                 // Copy actual to old
                 #statActualCommandOld := #statActualCommand;
                 #statModalCommandOld := #statModalCommand;

                 // Reset path data element and modal path data element
                 #statActualCommand := #statPathDataElementEmpty;
                 #statModalCommand := #statPathDataElementEmpty;

                 // Reset parameter counter for command
                 #statElementCounter := #statElementCounterEmpty;

                 // Initialize statCompletedPathDataCommand
                 #statActualCommand.pathDataElement := #statPathDataElementEmpty.pathDataElement;

                 FOR #tempCounter := 1 TO "LKINLANG_NUMBER_OF_CONDITIONS" DO
                   #statConditionsToCheck[#tempCounter] := #statConditionEmpty;
                   #statSetParametersInCmd[#tempCounter] := #statConditionEmpty;
                 END_FOR;

                 FOR #tempCounter := 1 TO "LKINLANG_MAX_NUMBER_OF_PARAMETERS_PER_LINE" DO
                   #tempParameterCounter[#tempCounter].parameterNumber := 0;
                   #tempParameterCounter[#tempCounter].counterValue := 0;
                 END_FOR;

                 // Save last positiong state (rel / abs)
                 #statPositioningModeOld := #statPositioningMode;

                 IF #statSearchedLine <= 0 THEN
                   // Next state --> Tokenize new line
                   #statStateIntern := #STATE_TOKENIZING;
                 ELSE
                   // Next state --> Search line
                   #statStateIntern := #STATE_SEARCH_LINE;
                 END_IF;

               END_IF;
             END_REGION RESET_AFTER_WRITE

             // ------------------------------------------------------------------------------------------
             // PreprocessingStop state for internal case
             // Switch to in case of preprocessingStop and do not execute other states
             // Wait until MovePath signalizes done
             // If done then go to STATE_TOKENIZING (continue with next line)
             // ------------------------------------------------------------------------------------------ 
             REGION PREPROCESSING_STOP
               // preprocessingStop State 
               IF #statStateIntern = #STATE_PREPROCESSING_STOP THEN
                 // preprocessingStop bit is set by parser and reset by MovePath 
                 // MovePath resets preprocessingStop if all commands are done
                 // Check if all commands are executed
                 IF #pathData.pointers.preprocessingStop = FALSE THEN
                   // Continue parsing
                   #statStateIntern := #STATE_TOKENIZING;
                 ELSE
                   ; // Stay here and wait
                 END_IF;
               END_IF;
             END_REGION PREPROCESSING_STOP

           END_FOR; // End of for loop 
         END_REGION FB_STATE_PARSING

         // ------------------------------------------------------------------------------------------
         // Error state for internal case
         // Switch to in case of error and do not execute other states
         // ------------------------------------------------------------------------------------------ 
         REGION ERROR_STATE
           // Error State 
           IF #statStateIntern = #STATE_ERROR THEN
             // Reset lineBuffer pointer
             #lineBuffer.pointers.retrievePointer := 0;
             #lineBuffer.pointers.addPointerRestarted := FALSE;
             IF #lineBuffer.pointers.endOfFile = FALSE THEN
               #lineBuffer.pointers.endOfFile := TRUE; // Signalize end to filehandler
             END_IF;
             // Reset file state
             IF #lineBuffer.info.fileState = "LKINLANG_FILE_STATE_RUNNING" THEN
               #lineBuffer.info.fileState := "LKINLANG_FILE_STATE_IDLE";
             END_IF;
           END_IF;
         END_REGION ERROR_STATE


         // ------------------------------------------------------------------------------------------
         // Stopping state in case stop input is triggered
         // Reset pointers where needed
         // ------------------------------------------------------------------------------------------ 
       #FB_STATE_STOPPING: // Stopping the parser
         REGION FB_STATE_STOPPING
           // Reset lineBuffer pointer
           #lineBuffer.pointers.retrievePointer := 0;

           // Reset pathData pointer 
           #pathData.pointers.addPointer := 0;
           #pathData.pointers.ignoreAddPointer := TRUE;
           #pathData.pointers.addPointerRestarted := FALSE;
           #pathData.pointers.bufferLocked := FALSE;
           #pathData.pointers.preprocessingStop := FALSE;

           // Set status
           #statStatus := #STATUS_COMMAND_ABORTED;
         END_REGION FB_STATE_STOPPING

       ELSE // Undefined state in state machine reached
         #statStatus := #ERR_UNDEFINED_STATE;
     END_CASE;

   END_REGION STATE_MACHINE


   REGION OUTPUTS
     // Write outputs
     IF (#statStatus = #STATUS_EXECUTION_FINISHED) AND (#statDone = FALSE) THEN // Execution finished without errors
       #statDone := TRUE;
       #statBusy := FALSE;
       #statCommandAborted := FALSE;
       #statError := FALSE;
       #statFBState := #FB_STATE_NO_PROCESSING; // Switch state machine to "no processing"

     ELSIF (#statStatus.%X15 = TRUE) AND (#statError = FALSE) THEN // Error occurred (#statStatus is 16#8000 to 16#FFFF)
       #statDone := FALSE;
       #statBusy := FALSE;
       #statCommandAborted := FALSE;
       #statError := TRUE;
       #statFBState := #FB_STATE_NO_PROCESSING; // Switch state machine to "no processing"

     ELSIF (#statStatus = #STATUS_COMMAND_ABORTED) AND (#statCommandAborted = FALSE) THEN // Commanded functionality has been aborted by another command
       #statDone := FALSE;
       #statBusy := FALSE;
       #statCommandAborted := TRUE;
       #statError := FALSE;
       #statFBState := #FB_STATE_NO_PROCESSING; // Switch state machine to "no processing"

     ELSIF (#tempExecute = FALSE) AND ((#statDone = TRUE) OR (#statError = TRUE) OR (#statCommandAborted = TRUE)) THEN // Reset outputs
       #statDone := FALSE;
       #statBusy := FALSE;
       #statCommandAborted := FALSE;
       #statError := FALSE;
       #statStatus := #STATUS_NO_CALL;
       // Reset application specific outputs
       #statErrorString := '';
       IF #lineBuffer.info.fileState = "LKINLANG_FILE_STATE_RUNNING" THEN
         #lineBuffer.info.fileState := "LKINLANG_FILE_STATE_IDLE";
       END_IF;
     END_IF;

     // Write static values to outputs
     #done := #statDone;
     #busy := #statBusy;
     #commandAborted := #statCommandAborted;
     #error := #statError;
     #status := #statStatus;
     #errorString := #statErrorString;
   END_REGION OUTPUTS


   //--------------------------------------------------------------------
   // End of Block LKinLang_Parser
   //--------------------------------------------------------------------
END_FUNCTION_BLOCK

FUNCTION_BLOCK "LKinLang_Filehandler"   // FB35451, SCL
TITLE = LKinLang_FileHandler
{ S7_Optimized_Access := 'TRUE' }
AUTHOR : tech.team.motioncontrol@siemens.com
FAMILY : LKinLang
VERSION : 1.1
// Transfer of data between memory card text file and PLC DB (buffer)
   VAR_INPUT
      executePlcToCard : Bool;   // Write data from buffer to card file
      executeCardToPlc : Bool;   // Write data from card file to buffer
      stop : Bool;   // stop the data transfer, abort the current command
      fileName : String;   // name of the card file (e.g. 'ProgramSlot.txt')
   END_VAR
   VAR_OUTPUT
      busy : Bool;   // TRUE: FB is not finished and new output values can be expected
      done : Bool;   // TRUE: Commanded action has been completed successfully
      dataTransferStopped : Bool;   // TRUE: The data transfer has been stopped
      error : Bool;   // Rising edge informs that an error occurred during the execution of
      status : Word := 16#7000;   // Current status of FB
      diagnostics : "LKinLang_typeFileHandlerDiagnostics";   // Diagnostics structure of FB
   END_VAR
   VAR_IN_OUT
      lineBuffer : "LKinLang_typeLineBuffer";   // String buffer connection
   END_VAR
   VAR
      statBusy : Bool;   // Static value for output busy
      statDone : Bool;   // Static value for output done
      statError : Bool;   // Static value for output error
      statCommandAborted : Bool;   // Static value for output commandAborted
      statPlcToCardOld : Bool;   // Old value of execute for edge detection
      statCardToPlcOld : Bool;   // Old value of execute for edge detection
      statStopOld : Bool;   // Old value of stop for edge detection
      statFBState : UInt;   // Static value for FB state
      statByteLine : Array[0..#NUMBER_OF_BYTES_PER_REQUEST] of Byte;   // Data storage for file read/write
      statByteLineCounter : UDInt;   // Counter/Index for the current byte line, which will be written with FileWriteC / Counter in the data storage
      statByteOffsetFile : UDInt;   // Offset for file read/write in the actual file on memory card / Offset for file read/write
      instFileWriteC : FileWriteC;
      instFileReadC : FileReadC;
      statLineCount : UDInt := 0;   // Actual line to write into the DB or into the file on the memory card / Number of lines from the current read file request
      statCurrentByteLine : Array[0..#NUMBER_OF_BYTES_PER_REQUEST] of Byte;   // Read bytes from actual read request
      statCharPosition : DInt;   // Conversion index CHAR-->STRING
      statBufferedLines : Array[0..#MAX_NUMBER_OF_LINES_PER_READ_REQUEST] of "LKinLang_typeLineContent";   // Buffer for single lines of file as string
      statLineIndex : DInt;   // Static store for last written line to continue FOR loop in case of exit
      statLineCountTotal : UDInt;   // Number of lines read in total
      statLastWrittenLine : UDInt;   // Static storing of the last written index
      statReadLineOld : UDInt;   // Static storing of the last read index
      statNumberOfRestBytes : UDInt;   // Number of bytes to be written on to the card
      statFileName : String;   // Static storing for the fileName input
      statFolderName : String := 'UserFiles';   // Static storing for the folderName
      statStatus : Word := 16#7000;   // Static value for output 'status'
      statSubfunctionStatus : Word;   // Static value for diagnostics subfunction status
      statLastLineWrite : UDInt;   // Static storing for the last written line
      statRequestedLine : UDInt;   // Static storing for requested line from pointer structure
      statOffset : UDInt;   // Static storing for the byte offset
   END_VAR
   VAR_TEMP
      tempExecutePlcToCard : Bool;   // Temporary value for input 'executePlcToCard'
      tempExecuteCardToPlc : Bool;   // Temporary value for input 'executeCardToPlc'
      tempStop : Bool;   // Temporary value for input 'stop'
      tempByteCounter : UDInt;   // Temporary byte counter
      tempLineCounter : DInt;   // Temporary line counter
      tempBufferIndex : DInt;   // Temporary index to write in lineBuffer
      tempCounter : DInt;   // Temporary general counter
      tempReadLineOld : UDInt;   // Temporary variable to store last read line
      tempRetrievePointer : DInt;   // Temporary variable for retrieve pointer
      tempEmptyByteLine : Array[0..#NUMBER_OF_BYTES_PER_REQUEST] of Byte;   // Temporary array to delete the byte line
      tempEmptyLine : "LKinLang_typeLineContent";   // Temporary line structure to delete a line
      tempEmptyDiagnostics : "LKinLang_typeFileHandlerDiagnostics";   // Empty diagnostics information (for initialization purposes only)
   END_VAR
   VAR CONSTANT
      MAX_NUMBER_OF_LINES_PER_READ_REQUEST : UDInt := 256;   // Maximum number of lines from one read request with FileReadC
      NUMBER_OF_BYTES_PER_REQUEST : UDInt := 256;   // Number of bytes for every read request with ReadFileC
      FB_STATE_NO_PROCESSING : UInt := 0;   // FB state: No processing
      FB_STATE_CARD_TO_PLC_INIT : UInt := 200;   // FB state: Card to PLC initialisation
      FB_STATE_CARD_TO_PLC_READ : UInt := 220;   // FB state: Card to PLC read data
      FB_STATE_CARD_TO_PLC_SEARCH_LINE : UInt := 240;   // FB state: Search specific line
      FB_STATE_CARD_TO_PLC_CONVERT : UInt := 250;   // FB state: Card to PLC convert byte to string
      FB_STATE_CARD_TO_PLC_WRITE_RING_BUFFER : UInt := 290;   // FB state: Card to PLC write string to buffer
      FB_STATE_PLC_TO_CARD_INIT : UInt := 300;   // FB state: PLC to Card initialisation
      FB_STATE_PLC_TO_CARD_READ : UInt := 320;   // FB state: PLC to Card convert string to byte
      FB_STATE_PLC_TO_CARD_WRITE : UInt := 350;   // FB state: PLC to Card write bytes to card
      FB_STATE_PLC_TO_CARD_READ_REST_BYTES : UInt := 360;   // FB state: PLC to Card get remaining bytes
      FB_STATE_PLC_TO_CARD_READ_REST_BYTES_RESULT : UInt := 370;   // FB state: PLC to Card evaluate remaining bytes
      FB_STATE_PLC_TO_CARD_DELETE_REST_BYTES : UInt := 380;   // FB state: PLC to Card delete remaining bytes
      FB_STATE_PLC_TO_CARD_DELETE_REST_BYTES_RESULT : UInt := 390;   // FB state: PLC to Card evaluate delete result
      STATUS_EXECUTION_FINISHED : Word := 16#0000;   // Execution finished without errors
      STATUS_NO_CALL : Word := 16#7000;   // No call of FB
      STATUS_FIRST_CALL : Word := 16#7001;   // First call of FB after enabling
      STATUS_SUBSEQUENT_CALL : Word := 16#7002;   // Subsequent call of FB
      STATUS_COMMAND_ABORTED : Word := 16#7FFF;   // Commanded functionality has been aborted by another command
      ERR_RETRIEVE_POINTER_INDEX : Word := 16#8001;   // Error due to retrieve pointer invalid
      ERR_INVALID_RETRIEVE_POINTER : Word := 16#8002;   // Index is outside of the range
      ERR_LINE_LENGTH : Word := 16#8004;   // Error due to line length being too low
      ERR_READ_AND_WRITE_CMD : Word := 16#8008;   // Error due to triggering both execute inputs
      ERR_UNDEFINED_STATE : Word := 16#8600;   // Error due to an undefined state in state machine
      ERR_READ_DATA_FROM_FILE : Word := 16#8601;   // Error due to FileReadC error
      ERR_WRITE_DATA_TO_FILE : Word := 16#8602;   // Error due to FileWriteC error
   END_VAR
BEGIN
   //=============================================================================
   // SIEMENS AG
   // (c)Copyright 2020 All Rights Reserved
   //-----------------------------------------------------------------------------
   // Library: LKinLang
   // Tested with: S7-1517T-3 PN/DP
   // Engineering: TIA Portal V15
   // Restrictions: ---
   // Requirements: S7-1500T FW 2.5
   // Functionality: LKinLang_FileHandler
   // Transfer of data between memory card text file and PLC DB (buffer)
   //
   // Support: tech.team.motioncontrol@siemens.com
   // Note: Parameter comments are only available in language 'English (United States)'
   //-----------------------------------------------------------------------------
   // Change log table:
   // Version      Date        Expert in charge    Changes applied
   // 01.00.00     28.05.2015  JW                  First created version
   // 01.00.01     15.11.2019  FR                  Added fileState info; dont write empty lines to card; Reset more statics in Init states
   // 01.01.00     23.03.2020  FR                  Added EndOfFile, Restart and requestedLine
   // 01.01.01     26.10.2020  FR                  Updated type conversions
   // 01.01.02     01.06.2021  FR                  Set "endOfFile" after saving
   //=============================================================================

   // Work with temporary value / create process image
   #tempExecutePlcToCard := #executePlcToCard;
   #tempExecuteCardToPlc := #executeCardToPlc;
   #tempStop := #stop;

   REGION TRIGGERING
     //===========================================================================================
     // check for rising edge of stop input
     // stop the current data transfer/command (when FB is busy and other/new data are required)
     IF (#tempStop = TRUE) AND (#statStopOld = FALSE) // And statBusy
     THEN
       // Perform stop procedure
       #statFBState := #FB_STATE_NO_PROCESSING;
       #statStatus := #STATUS_COMMAND_ABORTED;

       // if stop input is reset, new data transfers are possible, if stop is TRUE --> no data transfer
       //===========================================================================================
       // check for rising edge of one execute input
     ELSIF ((#tempExecutePlcToCard AND NOT #statPlcToCardOld) XOR (#tempExecuteCardToPlc AND NOT #statCardToPlcOld))
       AND (#statStatus = #STATUS_NO_CALL) // Triggering of new jobs during file transfer is not possible (stop required)
       AND (#tempStop = FALSE) // Stop input must be false
     THEN
       // FB triggered with one execute
       //-----------------------------------------------------------------------------------
       // First call; initialize FB
       #lineBuffer.pointers.endOfFile := FALSE;
       #statDone := FALSE;
       #statBusy := TRUE;
       #statError := FALSE;
       #statStatus := #STATUS_FIRST_CALL;

       // State machine - start processing depending on input
       IF #tempExecutePlcToCard THEN
         #statFBState := #FB_STATE_PLC_TO_CARD_INIT;
       ELSIF #tempExecuteCardToPlc THEN
         #statFBState := #FB_STATE_CARD_TO_PLC_INIT;
       END_IF;

       // Initialize functionality: reset of variables, diagnostics, etc.
       #diagnostics := #tempEmptyDiagnostics;
       #statSubfunctionStatus := 16#00;

       //===========================================================================================
       // reading and writing command cannot be executed at the same time --> error by user
     ELSIF ((#tempExecutePlcToCard AND NOT #statPlcToCardOld) AND (#tempExecuteCardToPlc AND NOT #statCardToPlcOld))
     THEN
       #statStatus := #ERR_READ_AND_WRITE_CMD;

       //===========================================================================================
       // Set correct status after first call
     ELSIF (#statStatus = #STATUS_FIRST_CALL) THEN
       #statStatus := #STATUS_SUBSEQUENT_CALL;

     ELSIF #lineBuffer.pointers.restart THEN
       #lineBuffer.pointers.restart := FALSE;
       #lineBuffer.pointers.endOfFile := FALSE;
       //-----------------------------------------------------------------------------------
       // First call; initialize FB
       #statDone := FALSE;
       #statBusy := TRUE;
       #statError := FALSE;
       #statStatus := #STATUS_FIRST_CALL;

       // State machine - start processing depending on input
       #statFBState := #FB_STATE_CARD_TO_PLC_INIT;

       // Initialize functionality: reset of variables, diagnostics, etc.
       #diagnostics := #tempEmptyDiagnostics;
       #statSubfunctionStatus := 16#00;

     END_IF;

     // save inputs for edge detection
     #statPlcToCardOld := #tempExecutePlcToCard;
     #statCardToPlcOld := #tempExecuteCardToPlc;
     #statStopOld := #tempStop;
   END_REGION TRIGGERING

   IF (#statStatus = #STATUS_NO_CALL) THEN // Nothing to do -> End here to reduce "system load"
     RETURN;
   END_IF;

   // Check inputs cyclic
   REGION CYCLIC_CHECK
     IF #lineBuffer.pointers.requestedLine <> 0
       AND #statFBState >= #FB_STATE_CARD_TO_PLC_INIT
       AND #instFileReadC.Busy = FALSE
     THEN
       #statRequestedLine := #lineBuffer.pointers.requestedLine;
       #lineBuffer.pointers.requestedLine := 0;
       #statFBState := #FB_STATE_CARD_TO_PLC_INIT;
     END_IF;

     // Check endOfFile
     IF #lineBuffer.pointers.endOfFile THEN
       #statStatus := #STATUS_EXECUTION_FINISHED;
       #statFBState := #FB_STATE_NO_PROCESSING;
       #lineBuffer.info.fileState := "LKINLANG_FILE_STATE_IDLE";
     END_IF;
   END_REGION CYCLIC_CHECK


   REGION STATE_MACHINE
     CASE #statFBState OF // State machine of FB
       #FB_STATE_NO_PROCESSING: // No processing active
         ;

         // ------------------------------------------------------------------------------  
         // Set the variables to initial state for WRITING to the CARD and go to next step  
         // ------------------------------------------------------------------------------  
       #FB_STATE_PLC_TO_CARD_INIT:
         REGION plc_to_card_init
           // initialize variables
           #statLineCount := INT_TO_UINT("LKINLANG_FIRST_INDEX_LINE_BUFFER");
           #statFBState := #FB_STATE_PLC_TO_CARD_READ;
           #statByteOffsetFile := 0;
           #statNumberOfRestBytes := 0;

           // Check if there are empty lines --> do not write them 
           #statLastLineWrite := INT_TO_UDINT("LKINLANG_LAST_INDEX_LINE_BUFFER");

           FOR #tempCounter := "LKINLANG_LAST_INDEX_LINE_BUFFER" TO "LKINLANG_FIRST_INDEX_LINE_BUFFER" BY -1 DO
             IF #lineBuffer.lines[#tempCounter].number = 0 AND #lineBuffer.lines[#tempCounter].content = '' THEN
               // Check next index
               CONTINUE;
             ELSE
               // Line with content found
               #statLastLineWrite := DINT_TO_UDINT(#tempCounter);
               EXIT;
             END_IF;
           END_FOR;

           // Reset statlineBuffer
           FOR #tempCounter := 0 TO UDINT_TO_DINT(#MAX_NUMBER_OF_LINES_PER_READ_REQUEST) DO
             #statBufferedLines[#tempCounter].content := '';
             #statBufferedLines[#tempCounter].number := 0;
           END_FOR;

           // Reset byte line
           // Reset current byte line
           FOR #tempCounter := 0 TO UDINT_TO_DINT(#NUMBER_OF_BYTES_PER_REQUEST) DO
             #statByteLine[#tempCounter] := 16#0;
             #statCurrentByteLine[#tempCounter] := 16#0;
           END_FOR;

           // Set file status
           #lineBuffer.info.fileState := "LKINLANG_FILE_STATE_SAVING";

           // Check if file name is given or has to be taken from file info
           IF #fileName <> '' THEN
             #statFileName := #fileName;
           ELSE
             #statFileName := #lineBuffer.info.fileName;
           END_IF;

           // Check if file name is viable
           IF #statFileName = '' THEN
             #statStatus := #ERR_WRITE_DATA_TO_FILE;
             ; // Error --> no name specified
           END_IF;


         END_REGION

         // ------------------------------------------------------------------------------  
         // Write strings (Program) from ascii slot to card
         // Translate strings from buffer to bytes (#statByteLine)
         // Calculate the needed byte size and trigger FileWriteC
         // ------------------------------------------------------------------------------    
       #FB_STATE_PLC_TO_CARD_READ:
         REGION plc_to_card_read
           // Translate string line in byte array
           #statByteLine := #tempEmptyByteLine;
           #statByteLineCounter := 0;

           // exit commands at the end of this loop
           WHILE
             // exit loop, when last line of buffer is reached
             (#statLineCount <= #statLastLineWrite)
             // exit loop when too many bytes/chars are included in the next line to write them with the next command
             // (statByteLine too small --> one more FileWrite execute required)
             // 2 for CR/LF (2 more bytes required)

           DO

             IF (2 + #statByteLineCounter + INT_TO_UDINT(LEN(IN := #lineBuffer.lines[#statLineCount].content)) <= #NUMBER_OF_BYTES_PER_REQUEST) THEN

               Strg_TO_Chars(Strg := #lineBuffer.lines[#statLineCount].content,
                             pChars := UDINT_TO_DINT(#statByteLineCounter),
                             Cnt => #tempByteCounter,
                             Chars := #statByteLine);

               #statByteLineCounter += #tempByteCounter;

               // If it is not the last line of the buffer, write CR/LF
               IF #statLineCount < #statLastLineWrite THEN
                 // Add CR/LF -> line break for file on card
                 #statByteLine[#statByteLineCounter] := 16#0D;
                 #statByteLineCounter += 1;
                 #statByteLine[#statByteLineCounter] := 16#0A;
                 #statByteLineCounter += 1;
                 // Calc length of byte array
                 #instFileWriteC.Length := #statByteLineCounter;
               ELSE
                 // Last line number from the buffer is reached no CR/LF -> no line break needed
                 // Set number of bytes, which have to be written for the FileWriteC instance
                 #instFileWriteC.Length := #statByteLineCounter;
               END_IF;

               // Go to next line in the buffer (while condition will check, whether the string in the line will fit into the byte line)
               #statLineCount += 1;
             ELSE
               EXIT;
             END_IF;

           END_WHILE;

           // write Inputs of File Write
           #instFileWriteC.REQ := True;
           #instFileWriteC.Offset := #statByteOffsetFile;
           #statFBState := #FB_STATE_PLC_TO_CARD_WRITE;

         END_REGION

         // ------------------------------------------------------------------------------  
         // Waiting for file writing done
         // Increment byte counter
         // If last index of slot is reached then go to #FB_STATE_PLC_TO_CARD_READ_REST_BYTES
         // Else go back to #FB_STATE_PLC_TO_CARD_READ
         // ------------------------------------------------------------------------------      
       #FB_STATE_PLC_TO_CARD_WRITE:
         REGION plc_to_card_write
           // Wait for written line
           IF #instFileWriteC.Done THEN
             // Calc new position for next line in byte stream
             #statByteOffsetFile += #instFileWriteC.ResultLength;

             // Go to next state
             IF #statLineCount > #statLastLineWrite AND NOT (#statStatus = #ERR_WRITE_DATA_TO_FILE) THEN
               // Delete remaining bytes from file afterwards
               #statFBState := #FB_STATE_PLC_TO_CARD_READ_REST_BYTES;
             ELSE
               // read the next line from the buffer
               #statFBState := #FB_STATE_PLC_TO_CARD_READ;
             END_IF;

           ELSE
             ; // Wait for writing
           END_IF;

           // Error occured in system function
           IF #instFileWriteC.Error THEN
             #diagnostics.subfunctionStatus := #instFileWriteC.Status;
             #statStatus := #ERR_WRITE_DATA_TO_FILE;
           ELSE
             ; // no error
           END_IF;



         END_REGION

         // ------------------------------------------------------------------------------  
         // Start read request to get remaining bytes in file after writing
         // Go to #FB_STATE_PLC_TO_CARD_READ_REST_BYTES_RESULT
         // ------------------------------------------------------------------------------    
       #FB_STATE_PLC_TO_CARD_READ_REST_BYTES:
         REGION plc_to_card_rest_bytes
           // read from the end of written bytes to the end of the file to read the number of remaining bytes which should be deleted
           #instFileReadC.REQ := TRUE;
           #instFileReadC.Offset := #statByteOffsetFile + #statNumberOfRestBytes;
           #instFileReadC.Length := #NUMBER_OF_BYTES_PER_REQUEST; // maximum for length
           #statFBState := #FB_STATE_PLC_TO_CARD_READ_REST_BYTES_RESULT;
         END_REGION

         // ------------------------------------------------------------------------------  
         // Check if fileRead is done 
         // If there are no rest bytes then execution is finished
         // If there are rest bytes then go to #FB_STATE_PLC_TO_CARD_DELETE_REST_BYTES to delete them
         // ------------------------------------------------------------------------------    
       #FB_STATE_PLC_TO_CARD_READ_REST_BYTES_RESULT:
         REGION plc_to_card_read_rest_bytes_result

           // Wait for read request
           IF #instFileReadC.Done THEN
             // count number of rest bytes
             #statNumberOfRestBytes += #instFileReadC.ResultLength;

             // no rest bytes in file --> PLC to CARD finished
             IF #statNumberOfRestBytes = 0 THEN
               // deleting finished // ram to card finished
               #statStatus := #STATUS_EXECUTION_FINISHED;
               #lineBuffer.info.fileState := "LKINLANG_FILE_STATE_IDLE";
               #lineBuffer.pointers.endOfFile := TRUE;
             ELSIF #instFileReadC.ResultLength < #NUMBER_OF_BYTES_PER_REQUEST
             THEN
               // Set offset for first filwWriteC to delete bytes 
               #instFileWriteC.Offset := #statByteOffsetFile;

               // end of the file found
               #statFBState := #FB_STATE_PLC_TO_CARD_DELETE_REST_BYTES;
             ELSE
               // new read request for data, because end of the file could not be found yet
               #statFBState := #FB_STATE_PLC_TO_CARD_READ_REST_BYTES;
             END_IF;
             ; // Wait for writing
           END_IF;

           // Error occured in system function
           IF #instFileReadC.Error THEN
             #statSubfunctionStatus := #instFileReadC.Status;
             #statStatus := #ERR_READ_DATA_FROM_FILE;
           ELSE
             ; // no error
           END_IF;

         END_REGION

         // ------------------------------------------------------------------------------  
         // Write NUL to delete content after written lines
         // ------------------------------------------------------------------------------    
       #FB_STATE_PLC_TO_CARD_DELETE_REST_BYTES:
         REGION plc_to_card_delete_rest_bytes
           // overwrite the rest bytes with NULL (ASCII 16#00)

           // add CR / LF at the start when writing
           #tempEmptyByteLine[0] := 16#0D;
           #tempEmptyByteLine[1] := 16#0A;
           // set all array elements to NULL
           #statByteLine := #tempEmptyByteLine;


           // start to overwrite the rest bytes with NULL (delete not possible)
           // do not write more bytes in one line than accepted!
           #instFileWriteC.REQ := TRUE;

           // FR 03.05.2019
           // Do not set offset here as instFileWriteC.ResultLength still has a value and can not be added here 
           //#instFileWriteC.Offset := #statByteCounterFile; //+ #instFileWriteC.ResultLength;

           #instFileWriteC.Length := LIMIT(MN := 0, IN := #statNumberOfRestBytes, MX := "LKINLANG_LENGTH_OF_ASCII_LINE_STRING");
           #statFBState := #FB_STATE_PLC_TO_CARD_DELETE_REST_BYTES_RESULT;
         END_REGION


         // ------------------------------------------------------------------------------  
         // Check if writing was successful 
         // If there are more bytes to delete go back to #FB_STATE_PLC_TO_CARD_DELETE_REST_BYTES
         // If all bytes were deleted then execution is finished
         // ------------------------------------------------------------------------------    
       #FB_STATE_PLC_TO_CARD_DELETE_REST_BYTES_RESULT:
         REGION plc_to_card_delete_rest_bytes_result

           // wait for successful writing NUL data
           IF #instFileWriteC.Done THEN
             #statNumberOfRestBytes -= #instFileWriteC.ResultLength;
             IF #statNumberOfRestBytes <= 0
             THEN
               // deleting finished // ram to card finished
               #statStatus := #STATUS_EXECUTION_FINISHED;
               #lineBuffer.info.fileState := "LKINLANG_FILE_STATE_IDLE";
               #lineBuffer.pointers.endOfFile := TRUE;
             ELSE
               // FR 02.05.2019
               // Increase offset after deleting
               #instFileWriteC.Offset += #instFileWriteC.ResultLength;

               // new read request for data, because end of the file could not be found yet
               #statFBState := #FB_STATE_PLC_TO_CARD_DELETE_REST_BYTES;
             END_IF;
             ; // Wait for writing
           END_IF;

           // Error occured in system function
           IF #instFileWriteC.Error THEN
             #statSubfunctionStatus := #instFileWriteC.Status;
             #statStatus := #ERR_WRITE_DATA_TO_FILE;
           ELSE
             ; // no error
           END_IF;

         END_REGION

         // ------------------------------------------------------------------------------  
         // Set the variables to initial state for READING from CARD and go to next step  
         // ------------------------------------------------------------------------------  
       #FB_STATE_CARD_TO_PLC_INIT:
         REGION card_to_plc_init
           #statByteOffsetFile := 0;
           #statCharPosition := 0;
           #statFBState := #FB_STATE_CARD_TO_PLC_READ;
           #statLineCountTotal := 0;
           #instFileReadC.Offset := 0;
           #statReadLineOld := 0;
           #instFileReadC.Length := #NUMBER_OF_BYTES_PER_REQUEST;
           #lineBuffer.pointers.addPointer := "LKINLANG_FIRST_INDEX_LINE_BUFFER";
           // Reset addPointerRestarted bit initially
           #lineBuffer.pointers.addPointerRestarted := FALSE;
           #lineBuffer.pointers.bufferLocked := TRUE;
           #lineBuffer.pointers.ignoreAddPointer := FALSE;
           #lineBuffer.pointers.endOfFile := FALSE;
           #statFileName := #fileName;
           #statLastWrittenLine := 0;
           #statLineCount := 0;

           #lineBuffer.info.fileName := #statFileName;
           #lineBuffer.info.fileState := "LKINLANG_FILE_STATE_LOADING";


           // reset the complete buffer, if a new data are requested
           FOR #tempCounter := "LKINLANG_FIRST_INDEX_LINE_BUFFER" TO "LKINLANG_LAST_INDEX_LINE_BUFFER" BY 1 DO
             #lineBuffer.lines[#tempCounter] := #tempEmptyLine;
           END_FOR;

           // Reset statlineBuffer
           FOR #tempCounter := 0 TO UDINT_TO_DINT(#MAX_NUMBER_OF_LINES_PER_READ_REQUEST) DO
             #statBufferedLines[#tempCounter].content := '';
             #statBufferedLines[#tempCounter].number := 0;
           END_FOR;

           // Reset byte line
           // Reset current byte line
           FOR #tempCounter := 0 TO UDINT_TO_DINT(#NUMBER_OF_BYTES_PER_REQUEST) DO
             #statByteLine[#tempCounter] := 16#0;
             #statCurrentByteLine[#tempCounter] := 16#0;
           END_FOR;
         END_REGION


         // ------------------------------------------------------------------------------  
         // Trigger FileRead and go to #FB_STATE_CARD_TO_PLC_CONVERT
         // ------------------------------------------------------------------------------   
       #FB_STATE_CARD_TO_PLC_READ:
         REGION card_to_plc_read
           ;// Read first line from file and write in byte array
           #instFileReadC.REQ := True;
           IF #statRequestedLine = 0 THEN
             #statFBState := #FB_STATE_CARD_TO_PLC_CONVERT;
           ELSE
             #statFBState := #FB_STATE_CARD_TO_PLC_SEARCH_LINE;
           END_IF;
         END_REGION card_to_plc_read

         // ------------------------------------------------------------------------------  
         // Search specific line and start reading from there
         // ------------------------------------------------------------------------------   
       #FB_STATE_CARD_TO_PLC_SEARCH_LINE:
         REGION card_to_plc_search_line
           IF #instFileReadC.Done
           THEN
             // Check if requested line is first line 
             // --> No offset needed
             IF #statRequestedLine = 1 THEN
               #statOffset := 0;
               #instFileReadC.Offset := 0;
               #statLineCountTotal := 0;
               #statRequestedLine := 0;
               #lineBuffer.pointers.retrievePointer := 0;
               #lineBuffer.pointers.addPointerRestarted := FALSE;
               #statFBState := #FB_STATE_CARD_TO_PLC_READ;
             ELSE
               // loop over all read bytes
               WHILE #tempByteCounter < #instFileReadC.ResultLength DO

                 IF (#statByteLine[#tempByteCounter] = 16#0D) // CR
                 THEN // end of line detected

                   // raise line counter
                   #statLineCount += 1;
                   #tempByteCounter += 2; // continue with reading next line / jump over CR (OD) LF (OA)

                 ELSE // go to next byte and write it into string of the current line
                   #tempByteCounter += 1;
                 END_IF;

                 // Check if line counter is one before requested line 
                 // --> Do not read requested line as we search the starting offset the requested line
                 // Yes: Exit while loop and restart reading with correct (found) offset
                 // No: The search continues
                 IF #statLineCount = #statRequestedLine - 1 THEN
                   #statOffset := #instFileReadC.Offset + #tempByteCounter;
                   #instFileReadC.Offset := #statOffset;
                   #statLineCountTotal := #statLineCount;
                   #statRequestedLine := 0;
                   #lineBuffer.pointers.retrievePointer := 0;
                   #lineBuffer.pointers.addPointerRestarted := FALSE;
                   #statFBState := #FB_STATE_CARD_TO_PLC_READ;
                   EXIT;
                 END_IF;

               END_WHILE;

               // If line was not found, restart reading with next offset
               IF #statLineCount <> #statRequestedLine - 1
                 AND #statRequestedLine > 0
               THEN
                 #instFileReadC.Offset += #instFileReadC.ResultLength;
                 #statFBState := #FB_STATE_CARD_TO_PLC_READ;
               END_IF;
             END_IF;


           ELSIF (#instFileReadC.Error)
           THEN
             #statStatus := #ERR_READ_DATA_FROM_FILE;
             #statSubfunctionStatus := #instFileReadC.Status;
           ELSE
             ; // FileRead not done and no error
             // --> FileRead still busy
           END_IF;
         END_REGION card_to_plc_search_line


         // ------------------------------------------------------------------------------  
         // Convert read byte array to internal string array 
         // Go to #FB_STATE_CARD_TO_PLC_WRITE_RING_BUFFER
         // ------------------------------------------------------------------------------
       #FB_STATE_CARD_TO_PLC_CONVERT:
         REGION card_to_plc_convert
           // Convert read byte array in string array
           // waiting for "done" and switch to next state is missing
           // all from read string are written into the string array element 0 - no line break detection

           IF #instFileReadC.Done
           THEN

             #statLineCount := 0;

             // loop over all read bytes
             WHILE #tempByteCounter < #instFileReadC.ResultLength DO

               IF (#statByteLine[#tempByteCounter] = 16#0D) // CR
               THEN // end of line detected

                 // raise line counter
                 #statLineCount += 1;

                 // write data to internal array of string
                 Chars_TO_Strg(Chars := #statCurrentByteLine,
                               pChars := 0,
                               Cnt := DINT_TO_UINT(#statCharPosition),
                               Strg => #statBufferedLines[#statLineCount - 1].content);

                 #statBufferedLines[#statLineCount - 1].number := #statLineCount + #statLineCountTotal;

                 #tempByteCounter += 2; // continue with reading next line / jump over CR (OD) LF (OA)

                 #statCharPosition := 0;
                 #statCurrentByteLine := #tempEmptyByteLine;

               ELSIF #statByteLine[#tempByteCounter] = 16#0A // if LF at the beginning of read bytes, go to next byte
               THEN
                 #tempByteCounter += 1;

               ELSIF #statByteLine[#tempByteCounter] = 16#00 THEN // dont regard empty bytes
                 #tempByteCounter += 1;
               ELSE // go to next byte and write it into string of the current line
                 #statCurrentByteLine[#statCharPosition] := #statByteLine[#tempByteCounter];
                 #statCharPosition += 1;
                 #tempByteCounter += 1;
               END_IF;

               IF #statCharPosition > "LKINLANG_LENGTH_OF_ASCII_LINE_STRING" THEN
                 #statStatus := #ERR_LINE_LENGTH;
                 EXIT; // Changed RETURN to EXIT; FR 23.05.2019
               END_IF;

             END_WHILE;

             IF #statStatus.%X15 = FALSE THEN // Added FR 23.05.2019: Skip in case of error
               IF #instFileReadC.ResultLength < #NUMBER_OF_BYTES_PER_REQUEST
               THEN
                 // if last bytes of file have been read - end of file reached
                 // #statInternalState := #STATE_IDLE;

                 // raise line counter
                 #statLineCount += 1;

                 // write last data to buffered Array of String 
                 Chars_TO_Strg(Chars := #statCurrentByteLine,
                               pChars := 0,
                               Cnt := DINT_TO_UINT(#statCharPosition),
                               Strg => #statBufferedLines[#statLineCount - 1].content);

                 #statBufferedLines[#statLineCount - 1].number := #statLineCount + #statLineCountTotal;
               END_IF;

               #statLineIndex := 0;

               #statFBState := #FB_STATE_CARD_TO_PLC_WRITE_RING_BUFFER;
             ELSE
               ; // Error already set --> do nothing 
             END_IF;


           ELSIF (#instFileReadC.Error)
           THEN
             #statStatus := #ERR_READ_DATA_FROM_FILE;
             #statSubfunctionStatus := #instFileReadC.Status;
           ELSE
             ; // FileRead not done and no erro
             // --> FileRead still busy
           END_IF;
         END_REGION

         // ------------------------------------------------------------------------------  
         // Write internal string array to buffer outside
         // If all strings were read then execution is finished
         // else go back to #FB_STATE_CARD_TO_PLC_READ
         // ------------------------------------------------------------------------------
       #FB_STATE_CARD_TO_PLC_WRITE_RING_BUFFER:
         REGION card_to_plc_write_ring_buffer

           IF #lineBuffer.pointers.retrievePointer = 0 THEN
             #tempRetrievePointer := 1;
           ELSE
             #tempRetrievePointer := #lineBuffer.pointers.retrievePointer;
           END_IF;

           // check retrieve pointer, if pointer outside the index limits of the array (buffer) --> user error
           IF #tempRetrievePointer < "LKINLANG_FIRST_INDEX_LINE_BUFFER" OR #tempRetrievePointer > "LKINLANG_LAST_INDEX_LINE_BUFFER" THEN
             #statStatus := #ERR_INVALID_RETRIEVE_POINTER;
             RETURN;

             // check if the last line number is higher than the actual one --> retrieve pointer overtook addPointer --> Error
           ELSIF #statReadLineOld > #lineBuffer.lines[#tempRetrievePointer].number
           THEN // last read line cannot be higher than last written line --> user error
             #statStatus := #ERR_RETRIEVE_POINTER_INDEX;
             RETURN;
           END_IF;

           // tempLineCount: Zählervariable innerhalb statBufferedStrings[]
           // statLineIndex: Merker für zuletzt geschriebene Zeile zum Fortsetzen bei Abbruch der FOR Schleife
           // sratLineCount: Anzahl an gelesenen Zeilen aus FileReadC Funktion
           // statLineCountTotal: Anzahl bisher gelesene Zeilen
           // tempBufferIndex: Index in LineBuffer 
           // statAddPointer: AddPointer in LineBuffer

           FOR #tempLineCounter := #statLineIndex TO UDINT_TO_DINT((#statLineCount - 1)) BY 1 DO
             // calculate the correct array index in the target buffer
             #tempBufferIndex := (#tempLineCounter + UDINT_TO_DINT(#statLineCountTotal)) MOD ("LKINLANG_LAST_INDEX_LINE_BUFFER" + 1 - "LKINLANG_FIRST_INDEX_LINE_BUFFER");
             #tempBufferIndex := "LKINLANG_FIRST_INDEX_LINE_BUFFER" + #tempBufferIndex;

             // check if new data can be written into the buffer or if Filehandler has to wait for raising retrievePointer
             IF (((#lineBuffer.pointers.retrievePointer <= #lineBuffer.pointers.addPointer)
               AND NOT #lineBuffer.pointers.addPointerRestarted
               AND NOT (#lineBuffer.pointers.addPointer = "LKINLANG_LAST_INDEX_LINE_BUFFER"
               AND #lineBuffer.pointers.retrievePointer <= 1))
               OR ((#lineBuffer.pointers.retrievePointer > #lineBuffer.pointers.addPointer + 1)
               AND #lineBuffer.pointers.addPointerRestarted)) THEN

               // write values into the target buffer
               #lineBuffer.lines[#tempBufferIndex] := #statBufferedLines[#tempLineCounter];
               // save last written line for output
               #statLastWrittenLine := #statBufferedLines[#tempLineCounter].number;
               // save target index if loop will be repeated
               #statLineIndex := #tempLineCounter;


               IF (#lineBuffer.pointers.addPointer = "LKINLANG_LAST_INDEX_LINE_BUFFER") AND (#tempBufferIndex = "LKINLANG_FIRST_INDEX_LINE_BUFFER")
               THEN
                 #lineBuffer.pointers.addPointerRestarted := TRUE;
               END_IF;

               // write last add index
               #lineBuffer.pointers.addPointer := #tempBufferIndex;
               // it is allowed to read data from buffer
               #lineBuffer.pointers.bufferLocked := FALSE;
             ELSE
               #statLineIndex := #tempLineCounter;
               // ring buffer --> wait for raising "lastReadLine" to push new values to the ring buffer
               EXIT; // do not write new values to the target buffer --> exit the for loop
             END_IF;
           END_FOR;

           // save last read line number to make a check in next cycle
           // temp because of reference --> call by value needed
           #tempReadLineOld := #lineBuffer.lines[#tempRetrievePointer].number;
           #statReadLineOld := #tempReadLineOld;

           // check if all lines from last read request are already written into the buffer
           IF #statLastWrittenLine >= #statLineCount + #statLineCountTotal
           THEN // all lines from last read request are written into the buffer
             IF #instFileReadC.ResultLength < #NUMBER_OF_BYTES_PER_REQUEST
             THEN // last lines from file are already written into buffer (file end reached)
               #statStatus := #STATUS_EXECUTION_FINISHED;
               #lineBuffer.pointers.endOfFile := TRUE;
               #lineBuffer.info.fileState := "LKINLANG_FILE_STATE_IDLE";
             ELSE // request new bytes from file
               #statFBState := #FB_STATE_CARD_TO_PLC_READ;
               #statLineCountTotal := #statLineCountTotal + #statLineCount;
               #instFileReadC.Offset += #NUMBER_OF_BYTES_PER_REQUEST;
             END_IF;
           ELSE // wait for raising "lastReadLine" to overwrite already read lines in buffer
             ; // do nothing - keep internal state
           END_IF;

         END_REGION


       ELSE // Undefined state in state machine reached
         #statStatus := #ERR_UNDEFINED_STATE;
     END_CASE;

   END_REGION STATE_MACHINE

   // Write translated string line in file on card
   // It is possible to write 32 KByte (32.768 Byte) in one cycle

   // call instance if FileWriteC 
   #instFileWriteC(// REQ:=
                   Name := CONCAT(IN1 := CONCAT(IN1 := #statFolderName, IN2 := '/'), IN2 := #statFileName),
                   // Offset := #statByteCounterFile,
                   // Length := #statByteCounter,
                   // Done=> ,
                   // Busy=> ,
                   // Error=> ,
                   // Status=> ,
                   // ResultLength=>,
                   Data := #statByteLine);

   // Reset REQ input
   #instFileWriteC.REQ := False;


   // Read file from card
   // It is possible to read a file with a maximum size of 16 MByte

   // call instance of FileReadC
   #instFileReadC(// REQ:= _bool_in_,
                  Name := CONCAT(IN1 := CONCAT(IN1 := #statFolderName, IN2 := '/'), IN2 := #statFileName),
                  // Offset:=_udint_in_,
                  // Length:=_udint_in_,
                  // Done=>_bool_out_,
                  // Busy=>_bool_out_,
                  // Error=>_bool_out_,
                  // Status=>_word_out_,
                  // ResultLength=>_udint_out_,
                  Data := #statByteLine);

   // Reset REQ input
   #instFileReadC.REQ := False;


   REGION OUTPUTS
     // Write outputs
     IF (#statStatus = #STATUS_EXECUTION_FINISHED) AND (#statDone = FALSE) THEN // Execution finished without errors
       #statDone := TRUE;
       #statBusy := FALSE;
       #statCommandAborted := FALSE;
       #statError := FALSE;
       #statFBState := #FB_STATE_NO_PROCESSING; // Switch state machine to "no processing"

     ELSIF (#statStatus.%X15 = TRUE) AND (#statError = FALSE) THEN // Error occurred (#statStatus is 16#8000 to 16#FFFF)
       #statDone := FALSE;
       #statBusy := FALSE;
       #statCommandAborted := FALSE;
       #statError := TRUE;
       // Write diagnostics
       #diagnostics.stateNumber := #statFBState;
       #diagnostics.status := #statStatus;
       #diagnostics.subfunctionStatus := #statSubfunctionStatus;

       // Set file state
       #lineBuffer.info.fileState := "LKINLANG_FILE_STATE_STOPPED";

       #statFBState := #FB_STATE_NO_PROCESSING; // Switch state machine to "no processing"